   1066: 'GCU_ALARM_WORD_05_BIT_10', class GCU Alarms, trigger "60_Alarm_Data_GCU_ALARM_WORD_05" bit 2
   1067: 'GCU_ALARM_WORD_05_BIT_11', class GCU Alarms, trigger "60_Alarm_Data_GCU_ALARM_WORD_05" bit 3
   1068: 'GCU_ALARM_WORD_05_BIT_12', class GCU Alarms, trigger "60_Alarm_Data_GCU_ALARM_WORD_05" bit 4
   1069: 'GCU_ALARM_WORD_05_BIT_13', class GCU Alarms, trigger "60_Alarm_Data_GCU_ALARM_WORD_05" bit 5
   1070: 'GCU_ALARM_WORD_05_BIT_14', class GCU Alarms, trigger "60_Alarm_Data_GCU_ALARM_WORD_05" bit 6
   1071: 'GCU_ALARM_WORD_05_BIT_15', class GCU Alarms, trigger "60_Alarm_Data_GCU_ALARM_WORD_05" bit 7
   1072: 'GCU_ALARM_WORD_05_BIT_0', class GCU Alarms, trigger "60_Alarm_Data_GCU_ALARM_WORD_05" bit 8
   1073: 'GCU_ALARM_WORD_05_BIT_1', class GCU Alarms, trigger "60_Alarm_Data_GCU_ALARM_WORD_05" bit 9
   1074: 'GCU_ALARM_WORD_05_BIT_2', class GCU Alarms, trigger "60_Alarm_Data_GCU_ALARM_WORD_05" bit 10
   1075: 'GCU_ALARM_WORD_05_BIT_3', class GCU Alarms, trigger "60_Alarm_Data_GCU_ALARM_WORD_05" bit 11
   1076: 'GCU_ALARM_WORD_05_BIT_4', class GCU Alarms, trigger "60_Alarm_Data_GCU_ALARM_WORD_05" bit 12
   1077: 'GCU_ALARM_WORD_05_BIT_5', class GCU Alarms, trigger "60_Alarm_Data_GCU_ALARM_WORD_05" bit 13
   1078: 'GCU_ALARM_WORD_05_BIT_6', class GCU Alarms, trigger "60_Alarm_Data_GCU_ALARM_WORD_05" bit 14
   1079: 'GCU_ALARM_WORD_05_BIT_7', class GCU Alarms, trigger "60_Alarm_Data_GCU_ALARM_WORD_05" bit 15
   1080: 'GCU_ALARM_WORD_06_BIT_8', class GCU Alarms, trigger "60_Alarm_Data_GCU_ALARM_WORD_06" bit 0
   1081: 'GCU_ALARM_WORD_06_BIT_9', class GCU Alarms, trigger "60_Alarm_Data_GCU_ALARM_WORD_06" bit 1
   1082: 'GCU_ALARM_WORD_06_BIT_10', class GCU Alarms, trigger "60_Alarm_Data_GCU_ALARM_WORD_06" bit 2
   1083: 'GCU_ALARM_WORD_06_BIT_11', class GCU Alarms, trigger "60_Alarm_Data_GCU_ALARM_WORD_06" bit 3
   1084: 'GCU_ALARM_WORD_06_BIT_12', class GCU Alarms, trigger "60_Alarm_Data_GCU_ALARM_WORD_06" bit 4
   1085: 'GCU_ALARM_WORD_06_BIT_13', class GCU Alarms, trigger "60_Alarm_Data_GCU_ALARM_WORD_06" bit 5
   1086: 'GCU_ALARM_WORD_06_BIT_14', class GCU Alarms, trigger "60_Alarm_Data_GCU_ALARM_WORD_06" bit 6
   1087: 'GCU_ALARM_WORD_06_BIT_15', class GCU Alarms, trigger "60_Alarm_Data_GCU_ALARM_WORD_06" bit 7
   1088: 'GCU_ALARM_WORD_06_BIT_0', class GCU Alarms, trigger "60_Alarm_Data_GCU_ALARM_WORD_06" bit 8
   1089: 'GCU_ALARM_WORD_06_BIT_1', class GCU Alarms, trigger "60_Alarm_Data_GCU_ALARM_WORD_06" bit 9
   1090: 'GCU_ALARM_WORD_06_BIT_2', class GCU Alarms, trigger "60_Alarm_Data_GCU_ALARM_WORD_06" bit 10
   1091: 'GCU_ALARM_WORD_06_BIT_3', class GCU Alarms, trigger "60_Alarm_Data_GCU_ALARM_WORD_06" bit 11
   1092: 'GCU_ALARM_WORD_06_BIT_4', class GCU Alarms, trigger "60_Alarm_Data_GCU_ALARM_WORD_06" bit 12
   1093: 'GCU_ALARM_WORD_06_BIT_5', class GCU Alarms, trigger "60_Alarm_Data_GCU_ALARM_WORD_06" bit 13
   1094: 'GCU_ALARM_WORD_06_BIT_6', class GCU Alarms, trigger "60_Alarm_Data_GCU_ALARM_WORD_06" bit 14
   1095: 'GCU_ALARM_WORD_06_BIT_7', class GCU Alarms, trigger "60_Alarm_Data_GCU_ALARM_WORD_06" bit 15
   1096: 'GCU_ALARM_WORD_07_BIT_8', class GCU Alarms, trigger "60_Alarm_Data_GCU_ALARM_WORD_07" bit 0
   1097: 'GCU_ALARM_WORD_07_BIT_9', class GCU Alarms, trigger "60_Alarm_Data_GCU_ALARM_WORD_07" bit 1
   1098: 'GCU_ALARM_WORD_07_BIT_10', class GCU Alarms, trigger "60_Alarm_Data_GCU_ALARM_WORD_07" bit 2
   1099: 'GCU_ALARM_WORD_07_BIT_11', class GCU Alarms, trigger "60_Alarm_Data_GCU_ALARM_WORD_07" bit 3
   1100: 'GCU_ALARM_WORD_07_BIT_12', class GCU Alarms, trigger "60_Alarm_Data_GCU_ALARM_WORD_07" bit 4
   1101: 'GCU_ALARM_WORD_07_BIT_13', class GCU Alarms, trigger "60_Alarm_Data_GCU_ALARM_WORD_07" bit 5
   1102: 'GCU_ALARM_WORD_07_BIT_14', class GCU Alarms, trigger "60_Alarm_Data_GCU_ALARM_WORD_07" bit 6
   1103: 'GCU_ALARM_WORD_07_BIT_15', class GCU Alarms, trigger "60_Alarm_Data_GCU_ALARM_WORD_07" bit 7
   1104: 'GCU_ALARM_WORD_07_BIT_0', class GCU Alarms, trigger "60_Alarm_Data_GCU_ALARM_WORD_07" bit 8
   1105: 'GCU_ALARM_WORD_07_BIT_1', class GCU Alarms, trigger "60_Alarm_Data_GCU_ALARM_WORD_07" bit 9
   1106: 'GCU_ALARM_WORD_07_BIT_2', class GCU Alarms, trigger "60_Alarm_Data_GCU_ALARM_WORD_07" bit 10
   1107: 'GCU_ALARM_WORD_07_BIT_3', class GCU Alarms, trigger "60_Alarm_Data_GCU_ALARM_WORD_07" bit 11
   1108: 'GCU_ALARM_WORD_07_BIT_4', class GCU Alarms, trigger "60_Alarm_Data_GCU_ALARM_WORD_07" bit 12
   1109: 'GCU_ALARM_WORD_07_BIT_5', class GCU Alarms, trigger "60_Alarm_Data_GCU_ALARM_WORD_07" bit 13
   1110: 'GCU_ALARM_WORD_07_BIT_6', class GCU Alarms, trigger "60_Alarm_Data_GCU_ALARM_WORD_07" bit 14
   1111: 'GCU_ALARM_WORD_07_BIT_7', class GCU Alarms, trigger "60_Alarm_Data_GCU_ALARM_WORD_07" bit 15
   1112: 'GCU_ALARM_WORD_08_BIT_8', class GCU Alarms, trigger "60_Alarm_Data_GCU_ALARM_WORD_08" bit 0
   1113: 'GCU_ALARM_WORD_08_BIT_9', class GCU Alarms, trigger "60_Alarm_Data_GCU_ALARM_WORD_08" bit 1
   1114: 'GCU_ALARM_WORD_08_BIT_10', class GCU Alarms, trigger "60_Alarm_Data_GCU_ALARM_WORD_08" bit 2
   1115: 'GCU_ALARM_WORD_08_BIT_11', class GCU Alarms, trigger "60_Alarm_Data_GCU_ALARM_WORD_08" bit 3
   1116: 'GCU_ALARM_WORD_08_BIT_12', class GCU Alarms, trigger "60_Alarm_Data_GCU_ALARM_WORD_08" bit 4
   1117: 'GCU_ALARM_WORD_08_BIT_13', class GCU Alarms, trigger "60_Alarm_Data_GCU_ALARM_WORD_08" bit 5
   1118: 'GCU_ALARM_WORD_08_BIT_14', class GCU Alarms, trigger "60_Alarm_Data_GCU_ALARM_WORD_08" bit 6
   1119: 'GCU_ALARM_WORD_08_BIT_15', class GCU Alarms, trigger "60_Alarm_Data_GCU_ALARM_WORD_08" bit 7
   1120: 'GCU_ALARM_WORD_08_BIT_0', class GCU Alarms, trigger "60_Alarm_Data_GCU_ALARM_WORD_08" bit 8
   1121: 'GCU_ALARM_WORD_08_BIT_1', class GCU Alarms, trigger "60_Alarm_Data_GCU_ALARM_WORD_08" bit 9
   1122: 'GCU_ALARM_WORD_08_BIT_2', class GCU Alarms, trigger "60_Alarm_Data_GCU_ALARM_WORD_08" bit 10
   1123: 'GCU_ALARM_WORD_08_BIT_3', class GCU Alarms, trigger "60_Alarm_Data_GCU_ALARM_WORD_08" bit 11
   1124: 'GCU_ALARM_WORD_08_BIT_4', class GCU Alarms, trigger "60_Alarm_Data_GCU_ALARM_WORD_08" bit 12
   1125: 'GCU_ALARM_WORD_08_BIT_5', class GCU Alarms, trigger "60_Alarm_Data_GCU_ALARM_WORD_08" bit 13
   1126: 'GCU_ALARM_WORD_08_BIT_6', class GCU Alarms, trigger "60_Alarm_Data_GCU_ALARM_WORD_08" bit 14
   1127: 'GCU_ALARM_WORD_08_BIT_7', class GCU Alarms, trigger "60_Alarm_Data_GCU_ALARM_WORD_08" bit 15
   1128: 'GCU_ALARM_WORD_09_BIT_8', class GCU Alarms, trigger "60_Alarm_Data_GCU_ALARM_WORD_09" bit 0
   1129: 'GCU_ALARM_WORD_09_BIT_9', class GCU Alarms, trigger "60_Alarm_Data_GCU_ALARM_WORD_09" bit 1
   1130: 'GCU_ALARM_WORD_09_BIT_10', class GCU Alarms, trigger "60_Alarm_Data_GCU_ALARM_WORD_09" bit 2
   1131: 'GCU_ALARM_WORD_09_BIT_11', class GCU Alarms, trigger "60_Alarm_Data_GCU_ALARM_WORD_09" bit 3
   1132: 'GCU_ALARM_WORD_09_BIT_12', class GCU Alarms, trigger "60_Alarm_Data_GCU_ALARM_WORD_09" bit 4
   1133: 'GCU_ALARM_WORD_09_BIT_13', class GCU Alarms, trigger "60_Alarm_Data_GCU_ALARM_WORD_09" bit 5
   1134: 'GCU_ALARM_WORD_09_BIT_14', class GCU Alarms, trigger "60_Alarm_Data_GCU_ALARM_WORD_09" bit 6
   1135: 'GCU_ALARM_WORD_09_BIT_15', class GCU Alarms, trigger "60_Alarm_Data_GCU_ALARM_WORD_09" bit 7
   1136: 'GCU_ALARM_WORD_09_BIT_0', class GCU Alarms, trigger "60_Alarm_Data_GCU_ALARM_WORD_09" bit 8
   1137: 'GCU_ALARM_WORD_09_BIT_1', class GCU Alarms, trigger "60_Alarm_Data_GCU_ALARM_WORD_09" bit 9
   1138: 'GCU_ALARM_WORD_09_BIT_2', class GCU Alarms, trigger "60_Alarm_Data_GCU_ALARM_WORD_09" bit 10
   1139: 'GCU_ALARM_WORD_09_BIT_3', class GCU Alarms, trigger "60_Alarm_Data_GCU_ALARM_WORD_09" bit 11
   1140: 'GCU_ALARM_WORD_09_BIT_4', class GCU Alarms, trigger "60_Alarm_Data_GCU_ALARM_WORD_09" bit 12
   1141: 'GCU_ALARM_WORD_09_BIT_5', class GCU Alarms, trigger "60_Alarm_Data_GCU_ALARM_WORD_09" bit 13
   1142: 'GCU_ALARM_WORD_09_BIT_6', class GCU Alarms, trigger "60_Alarm_Data_GCU_ALARM_WORD_09" bit 14
   1143: 'GCU_ALARM_WORD_09_BIT_7', class GCU Alarms, trigger "60_Alarm_Data_GCU_ALARM_WORD_09" bit 15
   1144: 'PIT-358 FRESH WATER INLET PRESSURE', class GCU Warnings, trigger "62_Warning_Data_GCU_WARNING_WORD_01" bit 0
   1145: 'GCU_WARNING_WORD_01_BIT_9', class GCU Warnings, trigger "62_Warning_Data_GCU_WARNING_WORD_01" bit 1
   1146: 'GCU_WARNING_WORD_01_BIT_10', class GCU Warnings, trigger "62_Warning_Data_GCU_WARNING_WORD_01" bit 2
   1147: 'GCU_WARNING_WORD_01_BIT_11', class GCU Warnings, trigger "62_Warning_Data_GCU_WARNING_WORD_01" bit 3
   1148: 'GCU_WARNING_WORD_01_BIT_12', class GCU Warnings, trigger "62_Warning_Data_GCU_WARNING_WORD_01" bit 4
   1149: 'GCU_WARNING_WORD_01_BIT_13', class GCU Warnings, trigger "62_Warning_Data_GCU_WARNING_WORD_01" bit 5
   1150: 'GCU_WARNING_WORD_01_BIT_14', class GCU Warnings, trigger "62_Warning_Data_GCU_WARNING_WORD_01" bit 6
   1151: 'GCU_WARNING_WORD_01_BIT_15', class GCU Warnings, trigger "62_Warning_Data_GCU_WARNING_WORD_01" bit 7
   1152: 'PIT-348 CSW PRESSURE - OUT OF RANGE', class GCU Warnings, trigger "62_Warning_Data_GCU_WARNING_WORD_01" bit 8
   1153: 'LIT-304 LIQUID LEVEL - OUT OF RANGE', class GCU Warnings, trigger "62_Warning_Data_GCU_WARNING_WORD_01" bit 9
   1154: 'TIT-406 GAS TO DECK (OUTLET) TEMP - OUT OF RANGE', class GCU Warnings, trigger "62_Warning_Data_GCU_WARNING_WORD_01" bit 10
   1155: 'TIT-408 FRESH WATER COOLING TEMP - OUT OF RANGE', class GCU Warnings, trigger "62_Warning_Data_GCU_WARNING_WORD_01" bit 11
   1156: 'TIT-002 PGC DISCHARGE (OUTLET) TEMP - OUT OF RANGE', class GCU Warnings, trigger "62_Warning_Data_GCU_WARNING_WORD_01" bit 12
   1157: 'PIT-002 PGC DISCHARGE (OUTLET) PRESSURE - OUT OF RANGE', class GCU Warnings, trigger "62_Warning_Data_GCU_WARNING_WORD_01" bit 13
   1158: 'PIT-353 RECIRCULATION FRESH WATER PRESSURE - OUT OF RANGE', class GCU Warnings, trigger "62_Warning_Data_GCU_WARNING_WORD_01" bit 14
   1159: 'PIT-416 GAS TO DECK PRESSURE - OUT OF RANGE', class GCU Warnings, trigger "62_Warning_Data_GCU_WARNING_WORD_01" bit 15
   1160: 'PIT-002 - HIGH', class GCU Warnings, trigger "62_Warning_Data_GCU_WARNING_WORD_02" bit 0
   1161: 'PIT-353 FRESH WATER COOLING TO GCU - LOW', class GCU Warnings, trigger "62_Warning_Data_GCU_WARNING_WORD_02" bit 1
   1162: 'PIT-353 FRESH WATER COOLING TO GCU - HIGH', class GCU Warnings, trigger "62_Warning_Data_GCU_WARNING_WORD_02" bit 2
   1163: 'PIT-416 PROCESS GAS TO DECK PRESSURE - LOW', class GCU Warnings, trigger "62_Warning_Data_GCU_WARNING_WORD_02" bit 3
   1164: 'PIT-416 PROCESS GAS TO DECK PRESSURE - HIGH', class GCU Warnings, trigger "62_Warning_Data_GCU_WARNING_WORD_02" bit 4
   1165: 'PIT-358 BOOSTER FRESH WATER FILL PRESSURE - LOW', class GCU Warnings, trigger "62_Warning_Data_GCU_WARNING_WORD_02" bit 5
   1166: 'PIT-358 BOOSTER FRESH WATER FILL PRESSURE - HIGH', class GCU Warnings, trigger "62_Warning_Data_GCU_WARNING_WORD_02" bit 6
   1167: 'FS-350 FRESH WATER COOLING FLOW SWITCH - LOW FLOW5', class GCU Warnings, trigger "62_Warning_Data_GCU_WARNING_WORD_02" bit 7
   1168: 'CHECK PIT-348 COOLING SEAWATER PRESSURE', class GCU Warnings, trigger "62_Warning_Data_GCU_WARNING_WORD_02" bit 8
   1169: 'CHECK PIT-348 LOW COOLING SEAWATER PRESSURE', class GCU Warnings, trigger "62_Warning_Data_GCU_WARNING_WORD_02" bit 9
   1170: 'CHECK PIT-348 HIGH COOLING SEAWATER PRESSURE', class GCU Warnings, trigger "62_Warning_Data_GCU_WARNING_WORD_02" bit 10
   1171: 'CHECK LIT-304 GCU TANK LEVEL - HIGH', class GCU Warnings, trigger "62_Warning_Data_GCU_WARNING_WORD_02" bit 11
   1172: 'LIT-304 GCU LIQUID LEVEL - LOW', class GCU Warnings, trigger "62_Warning_Data_GCU_WARNING_WORD_02" bit 12
   1173: 'TIT-406 PROCESS GAS TO DECK TEMPERATURE - HIGH TEMP', class GCU Warnings, trigger "62_Warning_Data_GCU_WARNING_WORD_02" bit 13
   1174: 'TIT-408 FRESH WATER COOLING TO GCU TEMPERATURE - HIGH TEMP', class GCU Warnings, trigger "62_Warning_Data_GCU_WARNING_WORD_02" bit 14
   1175: 'CHECK TIT-002 PGC DISCHARGE (OUTLET) TEMPERATURE', class GCU Warnings, trigger "62_Warning_Data_GCU_WARNING_WORD_02" bit 15
   1176: 'GCU_WARNING', class GCU Warnings, trigger "62_Warning_Data_GCU_WARNING_WORD_03" bit 0
   1177: 'GCU_WARNING', class GCU Warnings, trigger "62_Warning_Data_GCU_WARNING_WORD_03" bit 1
   1178: 'GCU_WARNING', class GCU Warnings, trigger "62_Warning_Data_GCU_WARNING_WORD_03" bit 2
   1179: 'GCU_WARNING', class GCU Warnings, trigger "62_Warning_Data_GCU_WARNING_WORD_03" bit 3
   1180: 'GCU_WARNING', class GCU Warnings, trigger "62_Warning_Data_GCU_WARNING_WORD_03" bit 4
   1181: 'GCU_WARNING', class GCU Warnings, trigger "62_Warning_Data_GCU_WARNING_WORD_03" bit 5
   1182: 'GCU_WARNING', class GCU Warnings, trigger "62_Warning_Data_GCU_WARNING_WORD_03" bit 6
   1183: 'GCU_WARNING', class GCU Warnings, trigger "62_Warning_Data_GCU_WARNING_WORD_03" bit 7
   1184: 'LS-303 GCU LIQUID LEVEL - LOW', class GCU Warnings, trigger "62_Warning_Data_GCU_WARNING_WORD_03" bit 8
   1185: 'GCU_WARNING_WORD_03_BIT_1', class GCU Warnings, trigger "62_Warning_Data_GCU_WARNING_WORD_03" bit 9
   1186: 'GCU E-400 - FAULT', class GCU Warnings, trigger "62_Warning_Data_GCU_WARNING_WORD_03" bit 10
   1187: 'TIT-408 FRESH WATER COOLING TO GCU TEMPERATURE - HIGH HIGH TEMP', class GCU Warnings, trigger "62_Warning_Data_GCU_WARNING_WORD_03" bit 11
   1188: 'TIT-406 PROCESS GAS TO DECK TEMPERATURE - HIGH HIGH TEMP', class GCU Warnings, trigger "62_Warning_Data_GCU_WARNING_WORD_03" bit 12
   1189: 'GCU_WARNING_WORD_03_BIT_5', class GCU Warnings, trigger "62_Warning_Data_GCU_WARNING_WORD_03" bit 13
   1190: 'GCU_WARNING_WORD_03_BIT_6', class GCU Warnings, trigger "62_Warning_Data_GCU_WARNING_WORD_03" bit 14
   1191: 'GCU_WARNING_WORD_03_BIT_7', class GCU Warnings, trigger "62_Warning_Data_GCU_WARNING_WORD_03" bit 15
   1192: 'GCU_WARNING_WORD_04_BIT_8', class GCU Warnings, trigger "62_Warning_Data_GCU_WARNING_WORD_04" bit 0
   1193: 'GCU_WARNING_WORD_04_BIT_9', class GCU Warnings, trigger "62_Warning_Data_GCU_WARNING_WORD_04" bit 1
   1194: 'GCU_WARNING_WORD_04_BIT_10', class GCU Warnings, trigger "62_Warning_Data_GCU_WARNING_WORD_04" bit 2
   1195: 'GCU_WARNING_WORD_04_BIT_11', class GCU Warnings, trigger "62_Warning_Data_GCU_WARNING_WORD_04" bit 3
   1196: 'GCU_WARNING_WORD_04_BIT_12', class GCU Warnings, trigger "62_Warning_Data_GCU_WARNING_WORD_04" bit 4
   1197: 'GCU_WARNING_WORD_04_BIT_13', class GCU Warnings, trigger "62_Warning_Data_GCU_WARNING_WORD_04" bit 5
   1198: 'GCU_WARNING_WORD_04_BIT_14', class GCU Warnings, trigger "62_Warning_Data_GCU_WARNING_WORD_04" bit 6
   1199: 'GCU_WARNING_WORD_04_BIT_15', class GCU Warnings, trigger "62_Warning_Data_GCU_WARNING_WORD_04" bit 7
   1200: 'GCU_WARNING_WORD_04_BIT_0', class GCU Warnings, trigger "62_Warning_Data_GCU_WARNING_WORD_04" bit 8
   1201: 'GCU_WARNING_WORD_04_BIT_1', class GCU Warnings, trigger "62_Warning_Data_GCU_WARNING_WORD_04" bit 9
   1202: 'GCU_WARNING_WORD_04_BIT_2', class GCU Warnings, trigger "62_Warning_Data_GCU_WARNING_WORD_04" bit 10
   1203: 'GCU_WARNING_WORD_04_BIT_3', class GCU Warnings, trigger "62_Warning_Data_GCU_WARNING_WORD_04" bit 11
   1204: 'GCU_WARNING_WORD_04_BIT_4', class GCU Warnings, trigger "62_Warning_Data_GCU_WARNING_WORD_04" bit 12
   1205: 'GCU_WARNING_WORD_04_BIT_5', class GCU Warnings, trigger "62_Warning_Data_GCU_WARNING_WORD_04" bit 13
   1206: 'GCU_WARNING_WORD_04_BIT_6', class GCU Warnings, trigger "62_Warning_Data_GCU_WARNING_WORD_04" bit 14
   1207: 'GCU_WARNING_WORD_04_BIT_7', class GCU Warnings, trigger "62_Warning_Data_GCU_WARNING_WORD_04" bit 15
   1208: 'GCU_WARNING_WORD_05_BIT_8', class GCU Warnings, trigger "62_Warning_Data_GCU_WARNING_WORD_05" bit 0
   1209: 'GCU_WARNING_WORD_05_BIT_9', class GCU Warnings, trigger "62_Warning_Data_GCU_WARNING_WORD_05" bit 1
   1210: 'GCU_WARNING_WORD_05_BIT_10', class GCU Warnings, trigger "62_Warning_Data_GCU_WARNING_WORD_05" bit 2
   1211: 'GCU_WARNING_WORD_05_BIT_11', class GCU Warnings, trigger "62_Warning_Data_GCU_WARNING_WORD_05" bit 3
   1212: 'GCU_WARNING_WORD_05_BIT_12', class GCU Warnings, trigger "62_Warning_Data_GCU_WARNING_WORD_05" bit 4
   1213: 'GCU_WARNING_WORD_05_BIT_13', class GCU Warnings, trigger "62_Warning_Data_GCU_WARNING_WORD_05" bit 5
   1214: 'GCU_WARNING_WORD_05_BIT_14', class GCU Warnings, trigger "62_Warning_Data_GCU_WARNING_WORD_05" bit 6
   1215: 'GCU_WARNING_WORD_05_BIT_15', class GCU Warnings, trigger "62_Warning_Data_GCU_WARNING_WORD_05" bit 7
   1216: 'GCU_WARNING_WORD_05_BIT_0', class GCU Warnings, trigger "62_Warning_Data_GCU_WARNING_WORD_05" bit 8
   1217: 'GCU_WARNING_WORD_05_BIT_1', class GCU Warnings, trigger "62_Warning_Data_GCU_WARNING_WORD_05" bit 9
   1218: 'GCU_WARNING_WORD_05_BIT_2', class GCU Warnings, trigger "62_Warning_Data_GCU_WARNING_WORD_05" bit 10
   1219: 'GCU_WARNING_WORD_05_BIT_3', class GCU Warnings, trigger "62_Warning_Data_GCU_WARNING_WORD_05" bit 11
   1220: 'GCU_WARNING_WORD_05_BIT_4', class GCU Warnings, trigger "62_Warning_Data_GCU_WARNING_WORD_05" bit 12
   1221: 'GCU_WARNING_WORD_05_BIT_5', class GCU Warnings, trigger "62_Warning_Data_GCU_WARNING_WORD_05" bit 13
   1222: 'GCU_WARNING_WORD_05_BIT_6', class GCU Warnings, trigger "62_Warning_Data_GCU_WARNING_WORD_05" bit 14
   1223: 'GCU_WARNING_WORD_05_BIT_7', class GCU Warnings, trigger "62_Warning_Data_GCU_WARNING_WORD_05" bit 15
   1224: 'GCU_WARNING_WORD_06_BIT_8', class GCU Warnings, trigger "62_Warning_Data_GCU_WARNING_WORD_06" bit 0
   1225: 'GCU_WARNING_WORD_06_BIT_9', class GCU Warnings, trigger "62_Warning_Data_GCU_WARNING_WORD_06" bit 1
   1226: 'GCU_WARNING_WORD_06_BIT_10', class GCU Warnings, trigger "62_Warning_Data_GCU_WARNING_WORD_06" bit 2
   1227: 'GCU_WARNING_WORD_06_BIT_11', class GCU Warnings, trigger "62_Warning_Data_GCU_WARNING_WORD_06" bit 3
   1228: 'GCU_WARNING_WORD_06_BIT_12', class GCU Warnings, trigger "62_Warning_Data_GCU_WARNING_WORD_06" bit 4
   1229: 'GCU_WARNING_WORD_06_BIT_13', class GCU Warnings, trigger "62_Warning_Data_GCU_WARNING_WORD_06" bit 5
   1230: 'GCU_WARNING_WORD_06_BIT_14', class GCU Warnings, trigger "62_Warning_Data_GCU_WARNING_WORD_06" bit 6
   1231: 'GCU_WARNING_WORD_06_BIT_15', class GCU Warnings, trigger "62_Warning_Data_GCU_WARNING_WORD_06" bit 7
   1232: 'GCU_WARNING_WORD_06_BIT_0', class GCU Warnings, trigger "62_Warning_Data_GCU_WARNING_WORD_06" bit 8
   1233: 'GCU_WARNING_WORD_06_BIT_1', class GCU Warnings, trigger "62_Warning_Data_GCU_WARNING_WORD_06" bit 9
   1234: 'GCU_WARNING_WORD_06_BIT_2', class GCU Warnings, trigger "62_Warning_Data_GCU_WARNING_WORD_06" bit 10
   1235: 'GCU_WARNING_WORD_06_BIT_3', class GCU Warnings, trigger "62_Warning_Data_GCU_WARNING_WORD_06" bit 11
   1236: 'GCU_WARNING_WORD_06_BIT_4', class GCU Warnings, trigger "62_Warning_Data_GCU_WARNING_WORD_06" bit 12
   1237: 'GCU_WARNING_WORD_06_BIT_5', class GCU Warnings, trigger "62_Warning_Data_GCU_WARNING_WORD_06" bit 13
   1238: 'GCU_WARNING_WORD_06_BIT_6', class GCU Warnings, trigger "62_Warning_Data_GCU_WARNING_WORD_06" bit 14
   1239: 'GCU_WARNING_WORD_06_BIT_7', class GCU Warnings, trigger "62_Warning_Data_GCU_WARNING_WORD_06" bit 15
   1240: 'GCU_WARNING_WORD_07_BIT_8', class GCU Warnings, trigger "62_Warning_Data_GCU_WARNING_WORD_07" bit 0
   1241: 'GCU_WARNING_WORD_07_BIT_9', class GCU Warnings, trigger "62_Warning_Data_GCU_WARNING_WORD_07" bit 1
   1242: 'GCU_WARNING_WORD_07_BIT_10', class GCU Warnings, trigger "62_Warning_Data_GCU_WARNING_WORD_07" bit 2
   1243: 'GCU_WARNING_WORD_07_BIT_11', class GCU Warnings, trigger "62_Warning_Data_GCU_WARNING_WORD_07" bit 3
   1244: 'GCU_WARNING_WORD_07_BIT_12', class GCU Warnings, trigger "62_Warning_Data_GCU_WARNING_WORD_07" bit 4
   1245: 'GCU_WARNING_WORD_07_BIT_13', class GCU Warnings, trigger "62_Warning_Data_GCU_WARNING_WORD_07" bit 5
   1246: 'GCU_WARNING_WORD_07_BIT_14', class GCU Warnings, trigger "62_Warning_Data_GCU_WARNING_WORD_07" bit 6
   1247: 'GCU_WARNING_WORD_07_BIT_15', class GCU Warnings, trigger "62_Warning_Data_GCU_WARNING_WORD_07" bit 7
   1248: 'GCU_WARNING_WORD_07_BIT_0', class GCU Warnings, trigger "62_Warning_Data_GCU_WARNING_WORD_07" bit 8
   1249: 'GCU_WARNING_WORD_07_BIT_1', class GCU Warnings, trigger "62_Warning_Data_GCU_WARNING_WORD_07" bit 9
   1250: 'GCU_WARNING_WORD_07_BIT_2', class GCU Warnings, trigger "62_Warning_Data_GCU_WARNING_WORD_07" bit 10
   1251: 'GCU_WARNING_WORD_07_BIT_3', class GCU Warnings, trigger "62_Warning_Data_GCU_WARNING_WORD_07" bit 11
   1252: 'GCU_WARNING_WORD_07_BIT_4', class GCU Warnings, trigger "62_Warning_Data_GCU_WARNING_WORD_07" bit 12
   1253: 'GCU_WARNING_WORD_07_BIT_5', class GCU Warnings, trigger "62_Warning_Data_GCU_WARNING_WORD_07" bit 13
   1254: 'GCU_WARNING_WORD_07_BIT_6', class GCU Warnings, trigger "62_Warning_Data_GCU_WARNING_WORD_07" bit 14
   1255: 'GCU_WARNING_WORD_07_BIT_7', class GCU Warnings, trigger "62_Warning_Data_GCU_WARNING_WORD_07" bit 15
   1256: 'GCU_WARNING_WORD_08_BIT_8', class GCU Warnings, trigger "62_Warning_Data_GCU_WARNING_WORD_08" bit 0
   1257: 'GCU_WARNING_WORD_08_BIT_9', class GCU Warnings, trigger "62_Warning_Data_GCU_WARNING_WORD_08" bit 1
   1258: 'GCU_WARNING_WORD_08_BIT_10', class GCU Warnings, trigger "62_Warning_Data_GCU_WARNING_WORD_08" bit 2
   1259: 'GCU_WARNING_WORD_08_BIT_11', class GCU Warnings, trigger "62_Warning_Data_GCU_WARNING_WORD_08" bit 3
   1260: 'GCU_WARNING_WORD_08_BIT_12', class GCU Warnings, trigger "62_Warning_Data_GCU_WARNING_WORD_08" bit 4
   1261: 'GCU_WARNING_WORD_08_BIT_13', class GCU Warnings, trigger "62_Warning_Data_GCU_WARNING_WORD_08" bit 5
   1262: 'GCU_WARNING_WORD_08_BIT_14', class GCU Warnings, trigger "62_Warning_Data_GCU_WARNING_WORD_08" bit 6
   1263: 'GCU_WARNING_WORD_08_BIT_15', class GCU Warnings, trigger "62_Warning_Data_GCU_WARNING_WORD_08" bit 7
   1264: 'GCU_WARNING_WORD_08_BIT_0', class GCU Warnings, trigger "62_Warning_Data_GCU_WARNING_WORD_08" bit 8
   1265: 'GCU_WARNING_WORD_08_BIT_1', class GCU Warnings, trigger "62_Warning_Data_GCU_WARNING_WORD_08" bit 9
   1266: 'GCU_WARNING_WORD_08_BIT_2', class GCU Warnings, trigger "62_Warning_Data_GCU_WARNING_WORD_08" bit 10
   1267: 'GCU_WARNING_WORD_08_BIT_3', class GCU Warnings, trigger "62_Warning_Data_GCU_WARNING_WORD_08" bit 11
   1268: 'GCU_WARNING_WORD_08_BIT_4', class GCU Warnings, trigger "62_Warning_Data_GCU_WARNING_WORD_08" bit 12
   1269: 'GCU_WARNING_WORD_08_BIT_5', class GCU Warnings, trigger "62_Warning_Data_GCU_WARNING_WORD_08" bit 13
   1270: 'GCU_WARNING_WORD_08_BIT_6', class GCU Warnings, trigger "62_Warning_Data_GCU_WARNING_WORD_08" bit 14
   1271: 'GCU_WARNING_WORD_08_BIT_7', class GCU Warnings, trigger "62_Warning_Data_GCU_WARNING_WORD_08" bit 15
   1272: 'GCU_WARNING_WORD_09_BIT_8', class GCU Warnings, trigger "62_Warning_Data_GCU_WARNING_WORD_09" bit 0
   1273: 'GCU_WARNING_WORD_09_BIT_9', class GCU Warnings, trigger "62_Warning_Data_GCU_WARNING_WORD_09" bit 1
   1274: 'GCU_WARNING_WORD_09_BIT_10', class GCU Warnings, trigger "62_Warning_Data_GCU_WARNING_WORD_09" bit 2
   1275: 'GCU_WARNING_WORD_09_BIT_11', class GCU Warnings, trigger "62_Warning_Data_GCU_WARNING_WORD_09" bit 3
   1276: 'GCU_WARNING_WORD_09_BIT_12', class GCU Warnings, trigger "62_Warning_Data_GCU_WARNING_WORD_09" bit 4
   1277: 'GCU_WARNING_WORD_09_BIT_13', class GCU Warnings, trigger "62_Warning_Data_GCU_WARNING_WORD_09" bit 5
   1278: 'GCU_WARNING_WORD_09_BIT_14', class GCU Warnings, trigger "62_Warning_Data_GCU_WARNING_WORD_09" bit 6
   1279: 'GCU_WARNING_WORD_09_BIT_15', class GCU Warnings, trigger "62_Warning_Data_GCU_WARNING_WORD_09" bit 7
   1280: 'GCU_WARNING_WORD_09_BIT_0', class GCU Warnings, trigger "62_Warning_Data_GCU_WARNING_WORD_09" bit 8
   1281: 'GCU_WARNING_WORD_09_BIT_1', class GCU Warnings, trigger "62_Warning_Data_GCU_WARNING_WORD_09" bit 9
   1282: 'GCU_WARNING_WORD_09_BIT_2', class GCU Warnings, trigger "62_Warning_Data_GCU_WARNING_WORD_09" bit 10
   1283: 'GCU_WARNING_WORD_09_BIT_3', class GCU Warnings, trigger "62_Warning_Data_GCU_WARNING_WORD_09" bit 11
   1284: 'GCU_WARNING_WORD_09_BIT_4', class GCU Warnings, trigger "62_Warning_Data_GCU_WARNING_WORD_09" bit 12
   1285: 'GCU_WARNING_WORD_09_BIT_5', class GCU Warnings, trigger "62_Warning_Data_GCU_WARNING_WORD_09" bit 13
   1286: 'GCU_WARNING_WORD_09_BIT_6', class GCU Warnings, trigger "62_Warning_Data_GCU_WARNING_WORD_09" bit 14
   1287: 'GCU_WARNING_WORD_09_BIT_7', class GCU Warnings, trigger "62_Warning_Data_GCU_WARNING_WORD_09" bit 15
   2032: 'PT415 RIO1 DECK IG PRESSURE LOW LOW', class Tank Control Alarms, trigger "2060_Alarm_Data_BTCS_ALARM_WORD_03" bit 0
   2033: '', class Tank Control Alarms, trigger "2060_Alarm_Data_BTCS_ALARM_WORD_03" bit 1
   2034: 'PT415 RIO1 DECK IG PRESSURE HGH HIGH', class Tank Control Alarms, trigger "2060_Alarm_Data_BTCS_ALARM_WORD_03" bit 2
   2035: 'PT415 RIO3 DECK IG PRESSURE LOW LOW', class Tank Control Alarms, trigger "2060_Alarm_Data_BTCS_ALARM_WORD_03" bit 3
   2036: 'PT415 RIO3 DECK IG PRESSURE HGH HIGH', class Tank Control Alarms, trigger "2060_Alarm_Data_BTCS_ALARM_WORD_03" bit 4
   2037: 'PT415 RIO4 DECK IG PRESSURE LOW LOW', class Tank Control Alarms, trigger "2060_Alarm_Data_BTCS_ALARM_WORD_03" bit 5
   2038: 'PT415 RIO4 DECK IG PRESSURE HGH HIGH', class Tank Control Alarms, trigger "2060_Alarm_Data_BTCS_ALARM_WORD_03" bit 6
   2039: '', class Tank Control Alarms, trigger "2060_Alarm_Data_BTCS_ALARM_WORD_03" bit 7
   2040: 'CV422 5 STARBOARD GAS to TANK VALVE FAULT', class Tank Control Alarms, trigger "2060_Alarm_Data_BTCS_ALARM_WORD_03" bit 8
   2041: 'CV422 6 PORT GAS to TANK VALVE FAULT', class Tank Control Alarms, trigger "2060_Alarm_Data_BTCS_ALARM_WORD_03" bit 9
   2042: 'CV422 6 STARBOARD GAS to TANK VALVE FAULT', class Tank Control Alarms, trigger "2060_Alarm_Data_BTCS_ALARM_WORD_03" bit 10
   2043: 'CV422 APT GAS to TANK VALVE FAULT', class Tank Control Alarms, trigger "2060_Alarm_Data_BTCS_ALARM_WORD_03" bit 11
   2044: '', class Tank Control Alarms, trigger "2060_Alarm_Data_BTCS_ALARM_WORD_03" bit 12
   2045: '', class Tank Control Alarms, trigger "2060_Alarm_Data_BTCS_ALARM_WORD_03" bit 13
   2046: '', class Tank Control Alarms, trigger "2060_Alarm_Data_BTCS_ALARM_WORD_03" bit 14
   2047: '', class Tank Control Alarms, trigger "2060_Alarm_Data_BTCS_ALARM_WORD_03" bit 15
   2048: '', class Tank Control Alarms, trigger "2060_Alarm_Data_BTCS_ALARM_WORD_04" bit 0
   2049: '', class Tank Control Alarms, trigger "2060_Alarm_Data_BTCS_ALARM_WORD_04" bit 1
   2050: '', class Tank Control Alarms, trigger "2060_Alarm_Data_BTCS_ALARM_WORD_04" bit 2
   2051: '', class Tank Control Alarms, trigger "2060_Alarm_Data_BTCS_ALARM_WORD_04" bit 3
   2052: '', class Tank Control Alarms, trigger "2060_Alarm_Data_BTCS_ALARM_WORD_04" bit 4
   2053: '', class Tank Control Alarms, trigger "2060_Alarm_Data_BTCS_ALARM_WORD_04" bit 5
   2054: '', class Tank Control Alarms, trigger "2060_Alarm_Data_BTCS_ALARM_WORD_04" bit 6
   2055: '', class Tank Control Alarms, trigger "2060_Alarm_Data_BTCS_ALARM_WORD_04" bit 7
   2056: 'PT415 RIO5 DECK IG PRESSURE LOW LOW', class Tank Control Alarms, trigger "2060_Alarm_Data_BTCS_ALARM_WORD_04" bit 8
   2057: 'PT415 RIO5 DECK IG PRESSURE HGH HIGH', class Tank Control Alarms, trigger "2060_Alarm_Data_BTCS_ALARM_WORD_04" bit 9
   2058: 'PT415 RIO6 DECK IG PRESSURE LOW LOW', class Tank Control Alarms, trigger "2060_Alarm_Data_BTCS_ALARM_WORD_04" bit 10
   2059: 'PT415 RIO6 DECK IG PRESSURE HGH HIGH', class Tank Control Alarms, trigger "2060_Alarm_Data_BTCS_ALARM_WORD_04" bit 11
   2060: 'PT415 RIO7 DECK IG PRESSURE LOW LOW', class Tank Control Alarms, trigger "2060_Alarm_Data_BTCS_ALARM_WORD_04" bit 12
   2061: 'PT415 RIO7 DECK IG PRESSURE HIGH HIGH', class Tank Control Alarms, trigger "2060_Alarm_Data_BTCS_ALARM_WORD_04" bit 13
   2062: '', class Tank Control Alarms, trigger "2060_Alarm_Data_BTCS_ALARM_WORD_04" bit 14
   2063: '', class Tank Control Alarms, trigger "2060_Alarm_Data_BTCS_ALARM_WORD_04" bit 15
   2064: 'CV422 3 PORT GAS to TANK VALVE FAULT', class Tank Control Alarms, trigger "2060_Alarm_Data_BTCS_ALARM_WORD_02" bit 3
   2065: 'CV421 1 STARBOARD GAS to TANK VALVE FAULT', class Tank Control Alarms, trigger "2060_Alarm_Data_BTCS_ALARM_WORD_02" bit 2
   2066: 'CV421 3 STARBOARD GAS to TANK VALVE FAULT', class Tank Control Alarms, trigger "2060_Alarm_Data_BTCS_ALARM_WORD_02" bit 4
   2067: 'CV422 5 PORT GAS to TANK VALVE FAULT', class Tank Control Alarms, trigger "2060_Alarm_Data_BTCS_ALARM_WORD_02" bit 7
   2068: 'CV421 4 STARBOARD GAS to TANK VALVE FAULT', class Tank Control Alarms, trigger "2060_Alarm_Data_BTCS_ALARM_WORD_02" bit 6
   2069: 'CV422 4 PORT GAS to TANK VALVE FAULT', class Tank Control Alarms, trigger "2060_Alarm_Data_BTCS_ALARM_WORD_02" bit 5
   2070: 'PS-436 2 BALLAST TANK PRESSURE - HIGH', class Tank Control Alarms, trigger "2060_Alarm_Data_BTCS_ALARM_WORD_01" bit 14
   2071: 'LS-425 2 STARBOARD LEVEL - HIGH HIGH', class Tank Control Alarms, trigger "2060_Alarm_Data_BTCS_ALARM_WORD_01" bit 13
   2072: 'LS-425 2 PORT LEVEL - HIGH HIGH', class Tank Control Alarms, trigger "2060_Alarm_Data_BTCS_ALARM_WORD_01" bit 12
   2073: '600-TX-433 APT O2 MONITOR - LOW', class Tank Control Alarms, trigger "2060_Alarm_Data_BTCS_ALARM_WORD_01" bit 15
   2074: 'CV422 1 PORT GAS to TANK VALVE FAULT', class Tank Control Alarms, trigger "2060_Alarm_Data_BTCS_ALARM_WORD_02" bit 1
   2075: 'CV422 FPT GAS to TANK VALVE FAULT', class Tank Control Alarms, trigger "2060_Alarm_Data_BTCS_ALARM_WORD_02" bit 0
   2076: 'PIT-424 2 STARBOARD TANK PRESSURE - HIGH HIGH', class Tank Control Alarms, trigger "2060_Alarm_Data_BTCS_ALARM_WORD_02" bit 15
   2077: 'PIT-424 2 STARBOARD TANK PRESSURE - LOW LOW', class Tank Control Alarms, trigger "2060_Alarm_Data_BTCS_ALARM_WORD_02" bit 14
   2078: 'PIT-415 2 STARBOARD DECK IG PRESSURE - LOW LOW', class Tank Control Alarms, trigger "2060_Alarm_Data_BTCS_ALARM_WORD_02" bit 10
   2079: 'PIT-415 2 PORT DECK IG PRESSURE - HIGH HIGH', class Tank Control Alarms, trigger "2060_Alarm_Data_BTCS_ALARM_WORD_02" bit 9
   2080: 'PIT-415 2 PORT DECK IG PRESSURE - LOW LOW', class Tank Control Alarms, trigger "2060_Alarm_Data_BTCS_ALARM_WORD_02" bit 8
   2081: 'PIT-415 2 STARBOARD DECK IG PRESSURE - HIGH HIGH', class Tank Control Alarms, trigger "2060_Alarm_Data_BTCS_ALARM_WORD_02" bit 11
   2082: 'PIT-424 2 PORT TANK PRESSURE - HIGH HIGH', class Tank Control Alarms, trigger "2060_Alarm_Data_BTCS_ALARM_WORD_02" bit 13
   2083: 'PIT-424 2 PORT TANK PRESSURE - LOW LOW', class Tank Control Alarms, trigger "2060_Alarm_Data_BTCS_ALARM_WORD_02" bit 12
   2084: 'FIT-418 2 PORT USD FLOW - LOW LOW', class Tank Control Alarms, trigger "2060_Alarm_Data_BTCS_ALARM_WORD_01" bit 0
   2085: 'CV-442 2 PORT GAS to TANK VALVE FAULT', class Tank Control Alarms, trigger "2060_Alarm_Data_BTCS_ALARM_WORD_01" bit 8
   2086: 'FIT-419 2 STARBOARD MBG FLOW - HIGH HIGH', class Tank Control Alarms, trigger "2060_Alarm_Data_BTCS_ALARM_WORD_01" bit 7
   2087: 'CV-441 2 STARBOARD GAS to TANK VALVE FAULT', class Tank Control Alarms, trigger "2060_Alarm_Data_BTCS_ALARM_WORD_01" bit 9
   2088: 'TIT-436 2 STARBOARD BWT TEMP - HIGH HIGH', class Tank Control Alarms, trigger "2060_Alarm_Data_BTCS_ALARM_WORD_01" bit 11
   2089: 'TIT-436 2 PORT BWT TEMP - HIGH HIGH', class Tank Control Alarms, trigger "2060_Alarm_Data_BTCS_ALARM_WORD_01" bit 10
   2090: 'FIT-419 2 STARBOARD MBG FLOW - LOW LOW', class Tank Control Alarms, trigger "2060_Alarm_Data_BTCS_ALARM_WORD_01" bit 6
   2091: 'FIT-420 2 PORT MBG FLOW - HIGH HIGH', class Tank Control Alarms, trigger "2060_Alarm_Data_BTCS_ALARM_WORD_01" bit 3
   2092: 'FIT-420 2 PORT MBG FLOW - LOW LOW', class Tank Control Alarms, trigger "2060_Alarm_Data_BTCS_ALARM_WORD_01" bit 2
   2093: 'FIT-418 2 PORT USD FLOW - HIGH HIGH', class Tank Control Alarms, trigger "2060_Alarm_Data_BTCS_ALARM_WORD_01" bit 1
   2094: 'FIT-417 2 STARBOARD USD FLOW - HIGH HIGH', class Tank Control Alarms, trigger "2060_Alarm_Data_BTCS_ALARM_WORD_01" bit 5
   2095: 'FIT-417 2 STARBOARD USD FLOW - LOW LOW', class Tank Control Alarms, trigger "2060_Alarm_Data_BTCS_ALARM_WORD_01" bit 4
   2128: 'FIT-418 2 PORT USD FLOW - LOW', class Tank Control Warnings, trigger "2062_Warning_Data_BTCS_WARNING_WORD_01" bit 0
   2129: 'FIT-418 2 PORT USD FLOW - HIGH', class Tank Control Warnings, trigger "2062_Warning_Data_BTCS_WARNING_WORD_01" bit 1
   2130: 'FIT-420 2 PORT MBG FLOW - LOW', class Tank Control Warnings, trigger "2062_Warning_Data_BTCS_WARNING_WORD_01" bit 2
   2131: 'FIT-420 2 PORT MBG FLOW - HIGH', class Tank Control Warnings, trigger "2062_Warning_Data_BTCS_WARNING_WORD_01" bit 3
   2132: 'FIT-417 2 STARBOARD USD FLOW - LOW', class Tank Control Warnings, trigger "2062_Warning_Data_BTCS_WARNING_WORD_01" bit 4
   2133: 'FIT-417 2 STARBOARD USD FLOW - HIGH', class Tank Control Warnings, trigger "2062_Warning_Data_BTCS_WARNING_WORD_01" bit 5
   2134: 'FIT-419 2 STARBOARD MBG FLOW - LOW', class Tank Control Warnings, trigger "2062_Warning_Data_BTCS_WARNING_WORD_01" bit 6
   2135: 'FIT-419 2 STARBOARD MBG FLOW - HIGH', class Tank Control Warnings, trigger "2062_Warning_Data_BTCS_WARNING_WORD_01" bit 7
   2136: '600-TX-433 APT O2 MONITOR - LOW', class Tank Control Warnings, trigger "2062_Warning_Data_BTCS_WARNING_WORD_01" bit 8
